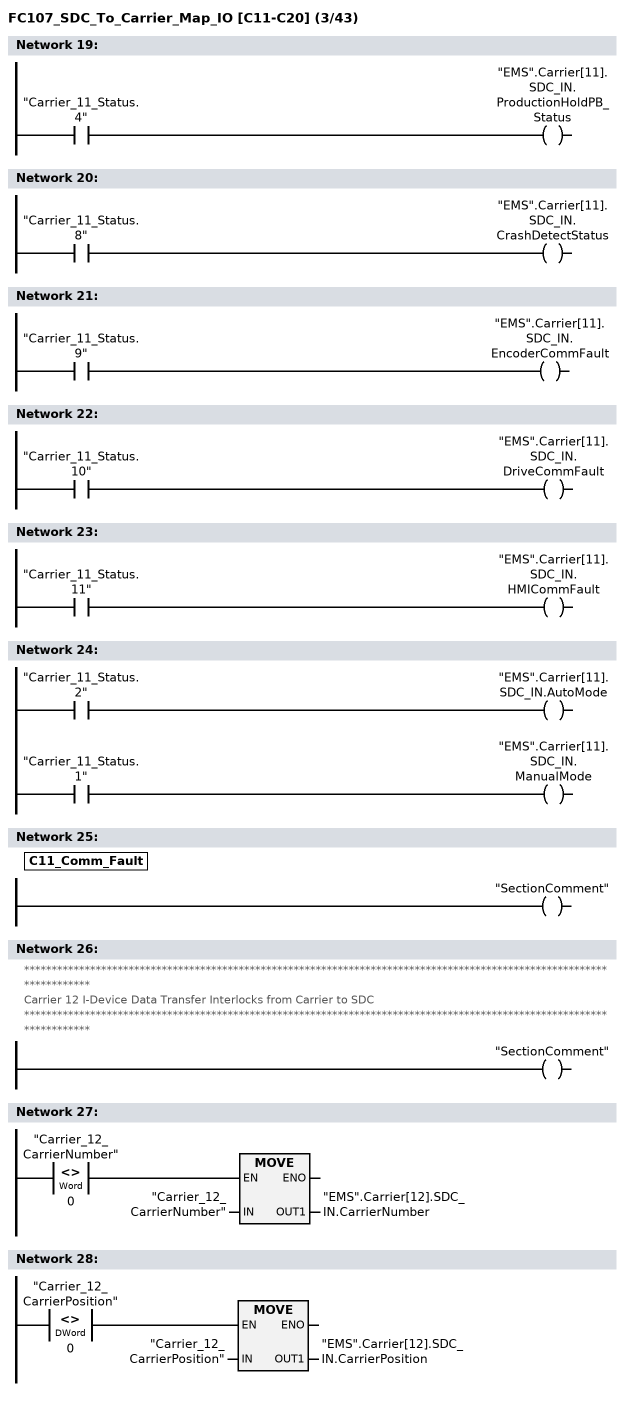
   RUNG wire#powerrail
      Contact( "Carrier_11_Status.4" )
      Coil( "EMS".Carrier[11].SDC_IN.ProductionHoldPB_Status )
   END_RUNG
   // the same network as SCL:
   "EMS".Carrier[11].SDC_IN.ProductionHoldPB_Status := "Carrier_11_Status.4";
END_REGION

REGION Network 20
   RUNG wire#powerrail
      Contact( "Carrier_11_Status.8" )
      Coil( "EMS".Carrier[11].SDC_IN.CrashDetectStatus )
   END_RUNG
   // the same network as SCL:
   "EMS".Carrier[11].SDC_IN.CrashDetectStatus := "Carrier_11_Status.8";
END_REGION

REGION Network 21
   RUNG wire#powerrail
      Contact( "Carrier_11_Status.9" )
      Coil( "EMS".Carrier[11].SDC_IN.EncoderCommFault )
   END_RUNG
   // the same network as SCL:
   "EMS".Carrier[11].SDC_IN.EncoderCommFault := "Carrier_11_Status.9";
END_REGION

REGION Network 22
   RUNG wire#powerrail
      Contact( "Carrier_11_Status.10" )
      Coil( "EMS".Carrier[11].SDC_IN.DriveCommFault )
   END_RUNG
   // the same network as SCL:
   "EMS".Carrier[11].SDC_IN.DriveCommFault := "Carrier_11_Status.10";
END_REGION

REGION Network 23
   RUNG wire#powerrail
      Contact( "Carrier_11_Status.11" )
      Coil( "EMS".Carrier[11].SDC_IN.HMICommFault )
   END_RUNG
   // the same network as SCL:
   "EMS".Carrier[11].SDC_IN.HMICommFault := "Carrier_11_Status.11";
END_REGION

REGION Network 24
   RUNG wire#powerrail
      Contact( "Carrier_11_Status.2" )
      Coil( "EMS".Carrier[11].SDC_IN.AutoMode )
   END_RUNG
   RUNG wire#powerrail
      Contact( "Carrier_11_Status.1" )
      Coil( "EMS".Carrier[11].SDC_IN.ManualMode )
   END_RUNG
   // the same network as SCL:
   "EMS".Carrier[11].SDC_IN.AutoMode := "Carrier_11_Status.2";
   "EMS".Carrier[11].SDC_IN.ManualMode := "Carrier_11_Status.1";
END_REGION

REGION Network 25
   Label( C11_Comm_Fault )
   RUNG wire#powerrail
      Coil( "SectionComment" )
   END_RUNG
   // the same network as SCL:
   C11_Comm_Fault:
   "SectionComment" := TRUE;
END_REGION

REGION Network 26
   // **********************************************************************************************************************
   // 
   // Carrier 12 I-Device Data Transfer Interlocks from Carrier to SDC
   // 
   // **********************************************************************************************************************
   RUNG wire#powerrail
      Coil( "SectionComment" )
   END_RUNG
   // the same network as SCL:
   "SectionComment" := TRUE;
END_REGION

REGION Network 27
   RUNG wire#powerrail
      { S7_Templates := "SrcType := Word" } NE_Contact(in1 := "Carrier_12_CarrierNumber", in2 := 0)
      Move(in := "Carrier_12_CarrierNumber", out1 => "EMS".Carrier[12].SDC_IN.CarrierNumber)
   END_RUNG
   // the same network as SCL:
   IF "Carrier_12_CarrierNumber" <> 0 THEN
       "EMS".Carrier[12].SDC_IN.CarrierNumber := "Carrier_12_CarrierNumber";
   END_IF;
END_REGION

REGION Network 28
   RUNG wire#powerrail
      { S7_Templates := "SrcType := DWord" } NE_Contact(in1 := "Carrier_12_CarrierPosition", in2 := 0)
      Move(in := "Carrier_12_CarrierPosition", out1 => "EMS".Carrier[12].SDC_IN.CarrierPosition)
   END_RUNG
   // the same network as SCL:
   IF "Carrier_12_CarrierPosition" <> 0 THEN
       "EMS".Carrier[12].SDC_IN.CarrierPosition := "Carrier_12_CarrierPosition";
   END_IF;
END_REGION

REGION Network 29
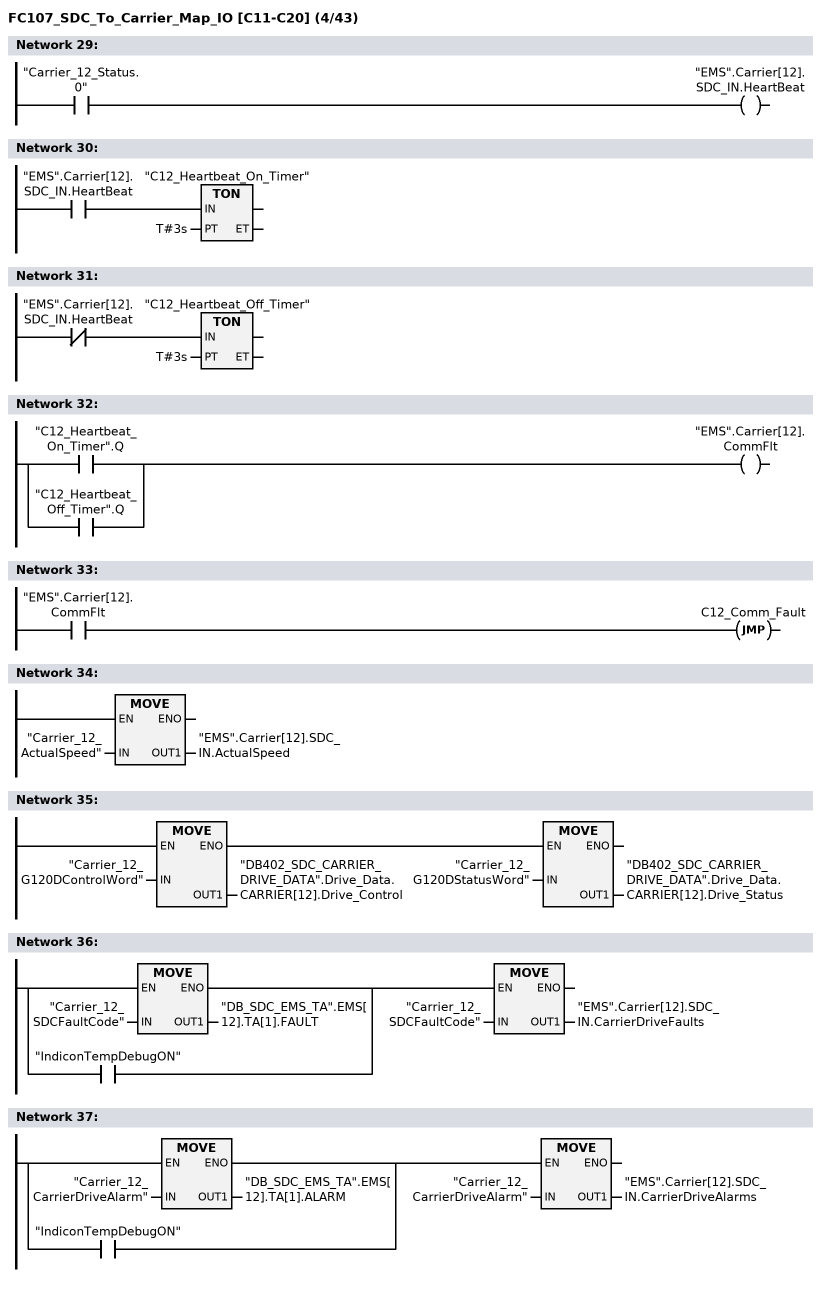
   RUNG wire#powerrail
      Contact( "Carrier_12_Status.0" )
      Coil( "EMS".Carrier[12].SDC_IN.HeartBeat )
   END_RUNG
   // the same network as SCL:
   "EMS".Carrier[12].SDC_IN.HeartBeat := "Carrier_12_Status.0";
END_REGION

REGION Network 30
   "C12_Heartbeat_On_Timer".TON(IN := "EMS".Carrier[12].SDC_IN.HeartBeat, PT := T#3s);
END_REGION

REGION Network 31
   "C12_Heartbeat_Off_Timer".TON(IN := NOT "EMS".Carrier[12].SDC_IN.HeartBeat, PT := T#3s);
END_REGION

REGION Network 32
   RUNG wire#powerrail
      Contact( "C12_Heartbeat_On_Timer".Q )
      wire#w1
      Coil( "EMS".Carrier[12].CommFlt )
   END_RUNG
   RUNG wire#powerrail
      Contact( "C12_Heartbeat_Off_Timer".Q )
   END_RUNG wire#w1
   // the same network as SCL:
   "EMS".Carrier[12].CommFlt := "C12_Heartbeat_On_Timer".Q OR "C12_Heartbeat_Off_Timer".Q;
END_REGION

REGION Network 33
   RUNG wire#powerrail
      Contact( "EMS".Carrier[12].CommFlt )
      JumpCoil( C12_Comm_Fault )
   END_RUNG
   // the same network as SCL:
   IF "EMS".Carrier[12].CommFlt THEN GOTO C12_Comm_Fault; END_IF;
END_REGION

REGION Network 34
   RUNG wire#powerrail
      Move(in := "Carrier_12_ActualSpeed", out1 => "EMS".Carrier[12].SDC_IN.ActualSpeed)
   END_RUNG
   // the same network as SCL:
   "EMS".Carrier[12].SDC_IN.ActualSpeed := "Carrier_12_ActualSpeed";
END_REGION

REGION Network 35
   RUNG wire#powerrail
      Move(in := "Carrier_12_G120DControlWord", out1 => "DB402_SDC_CARRIER_DRIVE_DATA".Drive_Data.CARRIER[12].Drive_Control)
      Move(in := "Carrier_12_G120DStatusWord", out1 => "DB402_SDC_CARRIER_DRIVE_DATA".Drive_Data.CARRIER[12].Drive_Status)
   END_RUNG
   // the same network as SCL:
   "DB402_SDC_CARRIER_DRIVE_DATA".Drive_Data.CARRIER[12].Drive_Control := "Carrier_12_G120DControlWord";
   "DB402_SDC_CARRIER_DRIVE_DATA".Drive_Data.CARRIER[12].Drive_Status := "Carrier_12_G120DStatusWord";
END_REGION

REGION Network 36
   RUNG wire#powerrail
      Move(in := "Carrier_12_SDCFaultCode", out1 => "DB_SDC_EMS_TA".EMS[12].TA[1].FAULT)
      wire#w1
      Move(in := "Carrier_12_SDCFaultCode", out1 => "EMS".Carrier[12].SDC_IN.CarrierDriveFaults)
   END_RUNG
   RUNG wire#powerrail
      Contact( "IndiconTempDebugON" )
   END_RUNG wire#w1
   // the same network as SCL:
   "DB_SDC_EMS_TA".EMS[12].TA[1].FAULT := "Carrier_12_SDCFaultCode";
   IF TRUE OR "IndiconTempDebugON" THEN
       "EMS".Carrier[12].SDC_IN.CarrierDriveFaults := "Carrier_12_SDCFaultCode";
   END_IF;
END_REGION

REGION Network 37
   RUNG wire#powerrail
      Move(in := "Carrier_12_CarrierDriveAlarm", out1 => "DB_SDC_EMS_TA".EMS[12].TA[1].ALARM)
      wire#w1
      Move(in := "Carrier_12_CarrierDriveAlarm", out1 => "EMS".Carrier[12].SDC_IN.CarrierDriveAlarms)
   END_RUNG
   RUNG wire#powerrail
      Contact( "IndiconTempDebugON" )
   END_RUNG wire#w1
   // the same network as SCL:
   "DB_SDC_EMS_TA".EMS[12].TA[1].ALARM := "Carrier_12_CarrierDriveAlarm";
   IF TRUE OR "IndiconTempDebugON" THEN
       "EMS".Carrier[12].SDC_IN.CarrierDriveAlarms := "Carrier_12_CarrierDriveAlarm";
   END_IF;
END_REGION

REGION Network 38
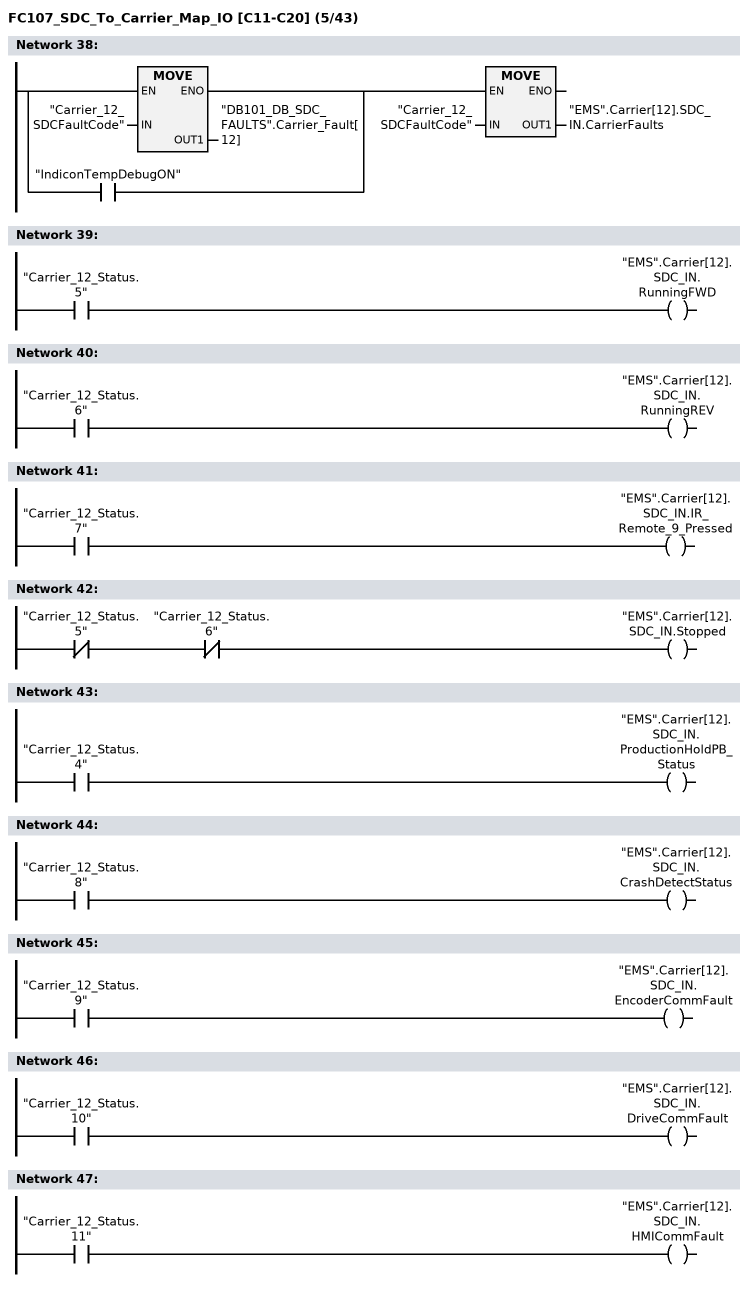
   RUNG wire#powerrail
      Move(in := "Carrier_12_SDCFaultCode", out1 => "DB101_DB_SDC_FAULTS".Carrier_Fault[12])
      wire#w1
      Move(in := "Carrier_12_SDCFaultCode", out1 => "EMS".Carrier[12].SDC_IN.CarrierFaults)
   END_RUNG
   RUNG wire#powerrail
      Contact( "IndiconTempDebugON" )
   END_RUNG wire#w1
   // the same network as SCL:
   "DB101_DB_SDC_FAULTS".Carrier_Fault[12] := "Carrier_12_SDCFaultCode";
   IF TRUE OR "IndiconTempDebugON" THEN
       "EMS".Carrier[12].SDC_IN.CarrierFaults := "Carrier_12_SDCFaultCode";
   END_IF;
END_REGION

REGION Network 39
   RUNG wire#powerrail
      Contact( "Carrier_12_Status.5" )
      Coil( "EMS".Carrier[12].SDC_IN.RunningFWD )
   END_RUNG
   // the same network as SCL:
   "EMS".Carrier[12].SDC_IN.RunningFWD := "Carrier_12_Status.5";
END_REGION

REGION Network 40
   RUNG wire#powerrail
      Contact( "Carrier_12_Status.6" )
      Coil( "EMS".Carrier[12].SDC_IN.RunningREV )
   END_RUNG
   // the same network as SCL:
   "EMS".Carrier[12].SDC_IN.RunningREV := "Carrier_12_Status.6";
END_REGION

REGION Network 41
   RUNG wire#powerrail
      Contact( "Carrier_12_Status.7" )
      Coil( "EMS".Carrier[12].SDC_IN.IR_Remote_9_Pressed )
   END_RUNG
   // the same network as SCL:
   "EMS".Carrier[12].SDC_IN.IR_Remote_9_Pressed := "Carrier_12_Status.7";
END_REGION

REGION Network 42
   RUNG wire#powerrail
      I_Contact( "Carrier_12_Status.5" )
      I_Contact( "Carrier_12_Status.6" )
      Coil( "EMS".Carrier[12].SDC_IN.Stopped )
   END_RUNG
   // the same network as SCL:
   "EMS".Carrier[12].SDC_IN.Stopped := NOT "Carrier_12_Status.5" AND NOT "Carrier_12_Status.6";
END_REGION

REGION Network 43
   RUNG wire#powerrail
      Contact( "Carrier_12_Status.4" )
      Coil( "EMS".Carrier[12].SDC_IN.ProductionHoldPB_Status )
   END_RUNG
   // the same network as SCL:
   "EMS".Carrier[12].SDC_IN.ProductionHoldPB_Status := "Carrier_12_Status.4";
END_REGION

REGION Network 44
   RUNG wire#powerrail
      Contact( "Carrier_12_Status.8" )
      Coil( "EMS".Carrier[12].SDC_IN.CrashDetectStatus )
   END_RUNG
   // the same network as SCL:
   "EMS".Carrier[12].SDC_IN.CrashDetectStatus := "Carrier_12_Status.8";
END_REGION

REGION Network 45
   RUNG wire#powerrail
      Contact( "Carrier_12_Status.9" )
      Coil( "EMS".Carrier[12].SDC_IN.EncoderCommFault )
   END_RUNG
   // the same network as SCL:
   "EMS".Carrier[12].SDC_IN.EncoderCommFault := "Carrier_12_Status.9";
END_REGION

REGION Network 46
   RUNG wire#powerrail
      Contact( "Carrier_12_Status.10" )
      Coil( "EMS".Carrier[12].SDC_IN.DriveCommFault )
   END_RUNG
   // the same network as SCL:
   "EMS".Carrier[12].SDC_IN.DriveCommFault := "Carrier_12_Status.10";
END_REGION

REGION Network 47
   RUNG wire#powerrail
      Contact( "Carrier_12_Status.11" )
      Coil( "EMS".Carrier[12].SDC_IN.HMICommFault )
   END_RUNG
   // the same network as SCL:
   "EMS".Carrier[12].SDC_IN.HMICommFault := "Carrier_12_Status.11";
END_REGION

REGION Network 48
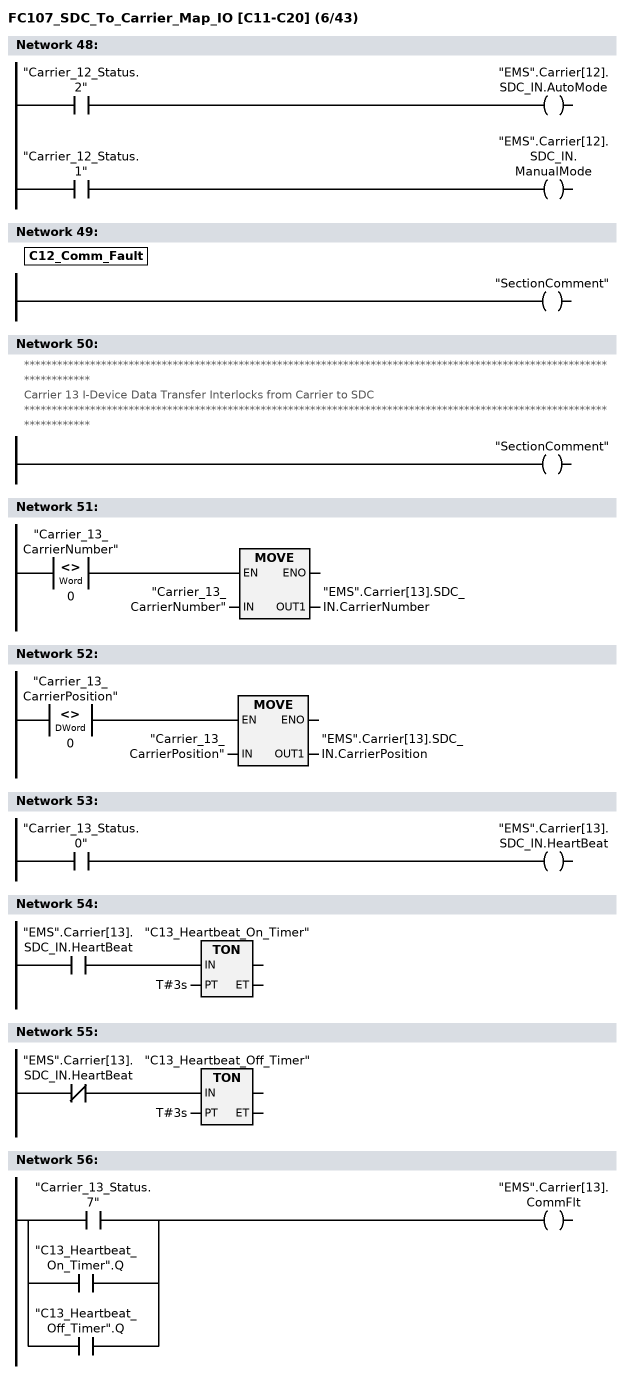
   RUNG wire#powerrail
      Contact( "Carrier_12_Status.2" )
      Coil( "EMS".Carrier[12].SDC_IN.AutoMode )
   END_RUNG
   RUNG wire#powerrail
      Contact( "Carrier_12_Status.1" )
      Coil( "EMS".Carrier[12].SDC_IN.ManualMode )
   END_RUNG
   // the same network as SCL:
   "EMS".Carrier[12].SDC_IN.AutoMode := "Carrier_12_Status.2";
   "EMS".Carrier[12].SDC_IN.ManualMode := "Carrier_12_Status.1";
END_REGION

REGION Network 49
   Label( C12_Comm_Fault )
   RUNG wire#powerrail
      Coil( "SectionComment" )
   END_RUNG
   // the same network as SCL:
   C12_Comm_Fault:
   "SectionComment" := TRUE;
END_REGION

REGION Network 50
   // **********************************************************************************************************************
   // 
   // Carrier 13 I-Device Data Transfer Interlocks from Carrier to SDC
   // 
   // **********************************************************************************************************************
   RUNG wire#powerrail
      Coil( "SectionComment" )
   END_RUNG
   // the same network as SCL:
   "SectionComment" := TRUE;
END_REGION

REGION Network 51
   RUNG wire#powerrail
      { S7_Templates := "SrcType := Word" } NE_Contact(in1 := "Carrier_13_CarrierNumber", in2 := 0)
      Move(in := "Carrier_13_CarrierNumber", out1 => "EMS".Carrier[13].SDC_IN.CarrierNumber)
   END_RUNG
   // the same network as SCL:
   IF "Carrier_13_CarrierNumber" <> 0 THEN
       "EMS".Carrier[13].SDC_IN.CarrierNumber := "Carrier_13_CarrierNumber";
   END_IF;
END_REGION

REGION Network 52
   RUNG wire#powerrail
      { S7_Templates := "SrcType := DWord" } NE_Contact(in1 := "Carrier_13_CarrierPosition", in2 := 0)
      Move(in := "Carrier_13_CarrierPosition", out1 => "EMS".Carrier[13].SDC_IN.CarrierPosition)
   END_RUNG
   // the same network as SCL:
   IF "Carrier_13_CarrierPosition" <> 0 THEN
       "EMS".Carrier[13].SDC_IN.CarrierPosition := "Carrier_13_CarrierPosition";
   END_IF;
END_REGION

REGION Network 53
   RUNG wire#powerrail
      Contact( "Carrier_13_Status.0" )
      Coil( "EMS".Carrier[13].SDC_IN.HeartBeat )
   END_RUNG
   // the same network as SCL:
   "EMS".Carrier[13].SDC_IN.HeartBeat := "Carrier_13_Status.0";
END_REGION

REGION Network 54
   "C13_Heartbeat_On_Timer".TON(IN := "EMS".Carrier[13].SDC_IN.HeartBeat, PT := T#3s);
END_REGION

REGION Network 55
   "C13_Heartbeat_Off_Timer".TON(IN := NOT "EMS".Carrier[13].SDC_IN.HeartBeat, PT := T#3s);
END_REGION

REGION Network 56
   RUNG wire#powerrail
      Contact( "Carrier_13_Status.7" )
      wire#w1
      Coil( "EMS".Carrier[13].CommFlt )
   END_RUNG
   RUNG wire#powerrail
      Contact( "C13_Heartbeat_On_Timer".Q )
   END_RUNG wire#w1
   RUNG wire#powerrail
      Contact( "C13_Heartbeat_Off_Timer".Q )
   END_RUNG wire#w1
   // the same network as SCL:
   "EMS".Carrier[13].CommFlt := "Carrier_13_Status.7" OR "C13_Heartbeat_On_Timer".Q OR "C13_Heartbeat_Off_Timer".Q;
END_REGION

REGION Network 57
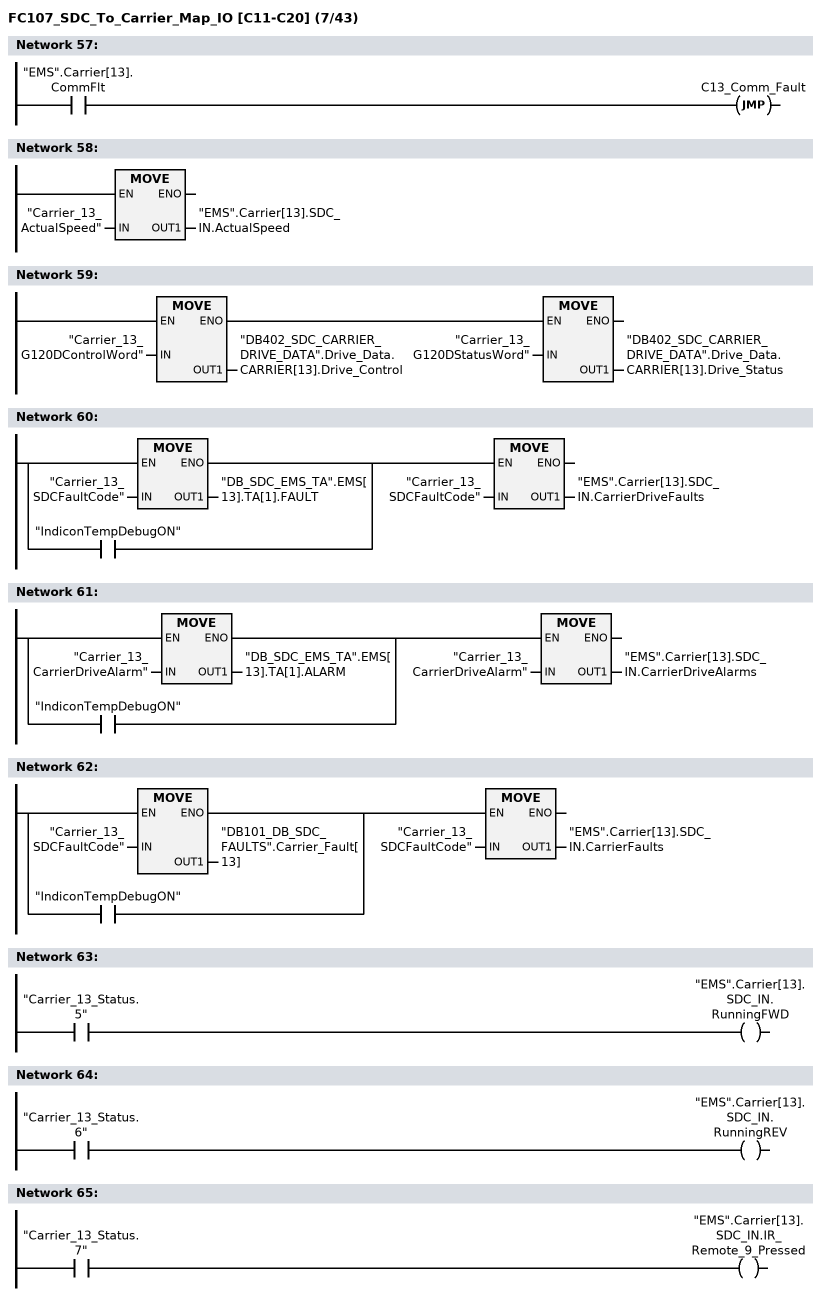
   RUNG wire#powerrail
      Contact( "EMS".Carrier[13].CommFlt )
      JumpCoil( C13_Comm_Fault )
   END_RUNG
   // the same network as SCL:
   IF "EMS".Carrier[13].CommFlt THEN GOTO C13_Comm_Fault; END_IF;
END_REGION

REGION Network 58
   RUNG wire#powerrail
      Move(in := "Carrier_13_ActualSpeed", out1 => "EMS".Carrier[13].SDC_IN.ActualSpeed)
   END_RUNG
   // the same network as SCL:
   "EMS".Carrier[13].SDC_IN.ActualSpeed := "Carrier_13_ActualSpeed";
END_REGION

REGION Network 59
   RUNG wire#powerrail
      Move(in := "Carrier_13_G120DControlWord", out1 => "DB402_SDC_CARRIER_DRIVE_DATA".Drive_Data.CARRIER[13].Drive_Control)
      Move(in := "Carrier_13_G120DStatusWord", out1 => "DB402_SDC_CARRIER_DRIVE_DATA".Drive_Data.CARRIER[13].Drive_Status)
   END_RUNG
   // the same network as SCL:
   "DB402_SDC_CARRIER_DRIVE_DATA".Drive_Data.CARRIER[13].Drive_Control := "Carrier_13_G120DControlWord";
   "DB402_SDC_CARRIER_DRIVE_DATA".Drive_Data.CARRIER[13].Drive_Status := "Carrier_13_G120DStatusWord";
END_REGION

REGION Network 60
   RUNG wire#powerrail
      Move(in := "Carrier_13_SDCFaultCode", out1 => "DB_SDC_EMS_TA".EMS[13].TA[1].FAULT)
      wire#w1
      Move(in := "Carrier_13_SDCFaultCode", out1 => "EMS".Carrier[13].SDC_IN.CarrierDriveFaults)
   END_RUNG
   RUNG wire#powerrail
      Contact( "IndiconTempDebugON" )
   END_RUNG wire#w1
   // the same network as SCL:
   "DB_SDC_EMS_TA".EMS[13].TA[1].FAULT := "Carrier_13_SDCFaultCode";
   IF TRUE OR "IndiconTempDebugON" THEN
       "EMS".Carrier[13].SDC_IN.CarrierDriveFaults := "Carrier_13_SDCFaultCode";
   END_IF;
END_REGION

REGION Network 61
   RUNG wire#powerrail
      Move(in := "Carrier_13_CarrierDriveAlarm", out1 => "DB_SDC_EMS_TA".EMS[13].TA[1].ALARM)
      wire#w1
      Move(in := "Carrier_13_CarrierDriveAlarm", out1 => "EMS".Carrier[13].SDC_IN.CarrierDriveAlarms)
   END_RUNG
   RUNG wire#powerrail
      Contact( "IndiconTempDebugON" )
   END_RUNG wire#w1
   // the same network as SCL:
   "DB_SDC_EMS_TA".EMS[13].TA[1].ALARM := "Carrier_13_CarrierDriveAlarm";
   IF TRUE OR "IndiconTempDebugON" THEN
       "EMS".Carrier[13].SDC_IN.CarrierDriveAlarms := "Carrier_13_CarrierDriveAlarm";
   END_IF;
END_REGION

REGION Network 62
   RUNG wire#powerrail
      Move(in := "Carrier_13_SDCFaultCode", out1 => "DB101_DB_SDC_FAULTS".Carrier_Fault[13])
      wire#w1
      Move(in := "Carrier_13_SDCFaultCode", out1 => "EMS".Carrier[13].SDC_IN.CarrierFaults)
   END_RUNG
   RUNG wire#powerrail
      Contact( "IndiconTempDebugON" )
   END_RUNG wire#w1
   // the same network as SCL:
   "DB101_DB_SDC_FAULTS".Carrier_Fault[13] := "Carrier_13_SDCFaultCode";
   IF TRUE OR "IndiconTempDebugON" THEN
       "EMS".Carrier[13].SDC_IN.CarrierFaults := "Carrier_13_SDCFaultCode";
   END_IF;
END_REGION

REGION Network 63
   RUNG wire#powerrail
      Contact( "Carrier_13_Status.5" )
      Coil( "EMS".Carrier[13].SDC_IN.RunningFWD )
   END_RUNG
   // the same network as SCL:
   "EMS".Carrier[13].SDC_IN.RunningFWD := "Carrier_13_Status.5";
END_REGION

REGION Network 64
   RUNG wire#powerrail
      Contact( "Carrier_13_Status.6" )
      Coil( "EMS".Carrier[13].SDC_IN.RunningREV )
   END_RUNG
   // the same network as SCL:
   "EMS".Carrier[13].SDC_IN.RunningREV := "Carrier_13_Status.6";
END_REGION

REGION Network 65
   RUNG wire#powerrail
      Contact( "Carrier_13_Status.7" )
      Coil( "EMS".Carrier[13].SDC_IN.IR_Remote_9_Pressed )
   END_RUNG
   // the same network as SCL:
   "EMS".Carrier[13].SDC_IN.IR_Remote_9_Pressed := "Carrier_13_Status.7";
END_REGION

REGION Network 66
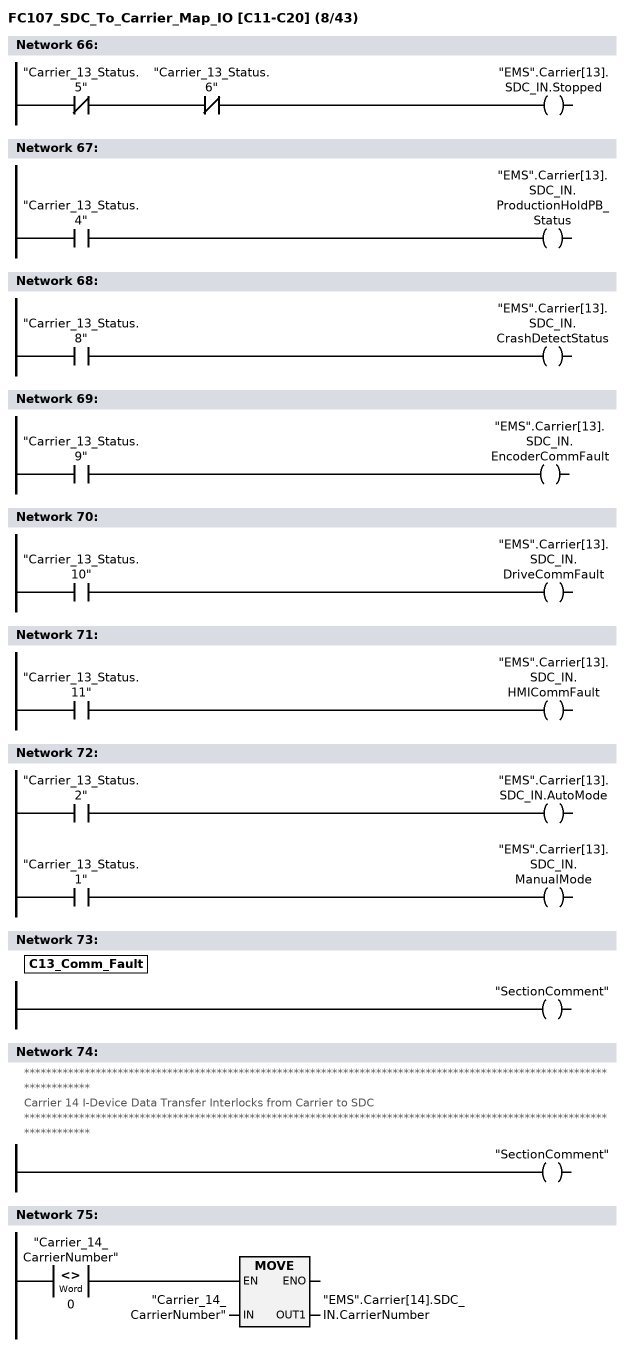
   RUNG wire#powerrail
      I_Contact( "Carrier_13_Status.5" )
      I_Contact( "Carrier_13_Status.6" )
      Coil( "EMS".Carrier[13].SDC_IN.Stopped )
   END_RUNG
   // the same network as SCL:
   "EMS".Carrier[13].SDC_IN.Stopped := NOT "Carrier_13_Status.5" AND NOT "Carrier_13_Status.6";
END_REGION

REGION Network 67
   RUNG wire#powerrail
      Contact( "Carrier_13_Status.4" )
      Coil( "EMS".Carrier[13].SDC_IN.ProductionHoldPB_Status )
   END_RUNG
   // the same network as SCL:
   "EMS".Carrier[13].SDC_IN.ProductionHoldPB_Status := "Carrier_13_Status.4";
END_REGION

REGION Network 68
   RUNG wire#powerrail
      Contact( "Carrier_13_Status.8" )
      Coil( "EMS".Carrier[13].SDC_IN.CrashDetectStatus )
   END_RUNG
   // the same network as SCL:
   "EMS".Carrier[13].SDC_IN.CrashDetectStatus := "Carrier_13_Status.8";
END_REGION

REGION Network 69
   RUNG wire#powerrail
      Contact( "Carrier_13_Status.9" )
      Coil( "EMS".Carrier[13].SDC_IN.EncoderCommFault )
   END_RUNG
   // the same network as SCL:
   "EMS".Carrier[13].SDC_IN.EncoderCommFault := "Carrier_13_Status.9";
END_REGION

REGION Network 70
   RUNG wire#powerrail
      Contact( "Carrier_13_Status.10" )
      Coil( "EMS".Carrier[13].SDC_IN.DriveCommFault )
   END_RUNG
   // the same network as SCL:
   "EMS".Carrier[13].SDC_IN.DriveCommFault := "Carrier_13_Status.10";
END_REGION

REGION Network 71
   RUNG wire#powerrail
      Contact( "Carrier_13_Status.11" )
      Coil( "EMS".Carrier[13].SDC_IN.HMICommFault )
   END_RUNG
   // the same network as SCL:
   "EMS".Carrier[13].SDC_IN.HMICommFault := "Carrier_13_Status.11";
END_REGION

REGION Network 72
   RUNG wire#powerrail
      Contact( "Carrier_13_Status.2" )
      Coil( "EMS".Carrier[13].SDC_IN.AutoMode )
   END_RUNG
   RUNG wire#powerrail
      Contact( "Carrier_13_Status.1" )
      Coil( "EMS".Carrier[13].SDC_IN.ManualMode )
   END_RUNG
   // the same network as SCL:
   "EMS".Carrier[13].SDC_IN.AutoMode := "Carrier_13_Status.2";
   "EMS".Carrier[13].SDC_IN.ManualMode := "Carrier_13_Status.1";
END_REGION

REGION Network 73
   Label( C13_Comm_Fault )
   RUNG wire#powerrail
      Coil( "SectionComment" )
   END_RUNG
   // the same network as SCL:
   C13_Comm_Fault:
   "SectionComment" := TRUE;
END_REGION

REGION Network 74
   // **********************************************************************************************************************
   // 
   // Carrier 14 I-Device Data Transfer Interlocks from Carrier to SDC
   // 
   // **********************************************************************************************************************
   RUNG wire#powerrail
      Coil( "SectionComment" )
   END_RUNG
   // the same network as SCL:
   "SectionComment" := TRUE;
END_REGION

REGION Network 75
   RUNG wire#powerrail
      { S7_Templates := "SrcType := Word" } NE_Contact(in1 := "Carrier_14_CarrierNumber", in2 := 0)
      Move(in := "Carrier_14_CarrierNumber", out1 => "EMS".Carrier[14].SDC_IN.CarrierNumber)
   END_RUNG
   // the same network as SCL:
   IF "Carrier_14_CarrierNumber" <> 0 THEN
       "EMS".Carrier[14].SDC_IN.CarrierNumber := "Carrier_14_CarrierNumber";
   END_IF;
END_REGION

REGION Network 76
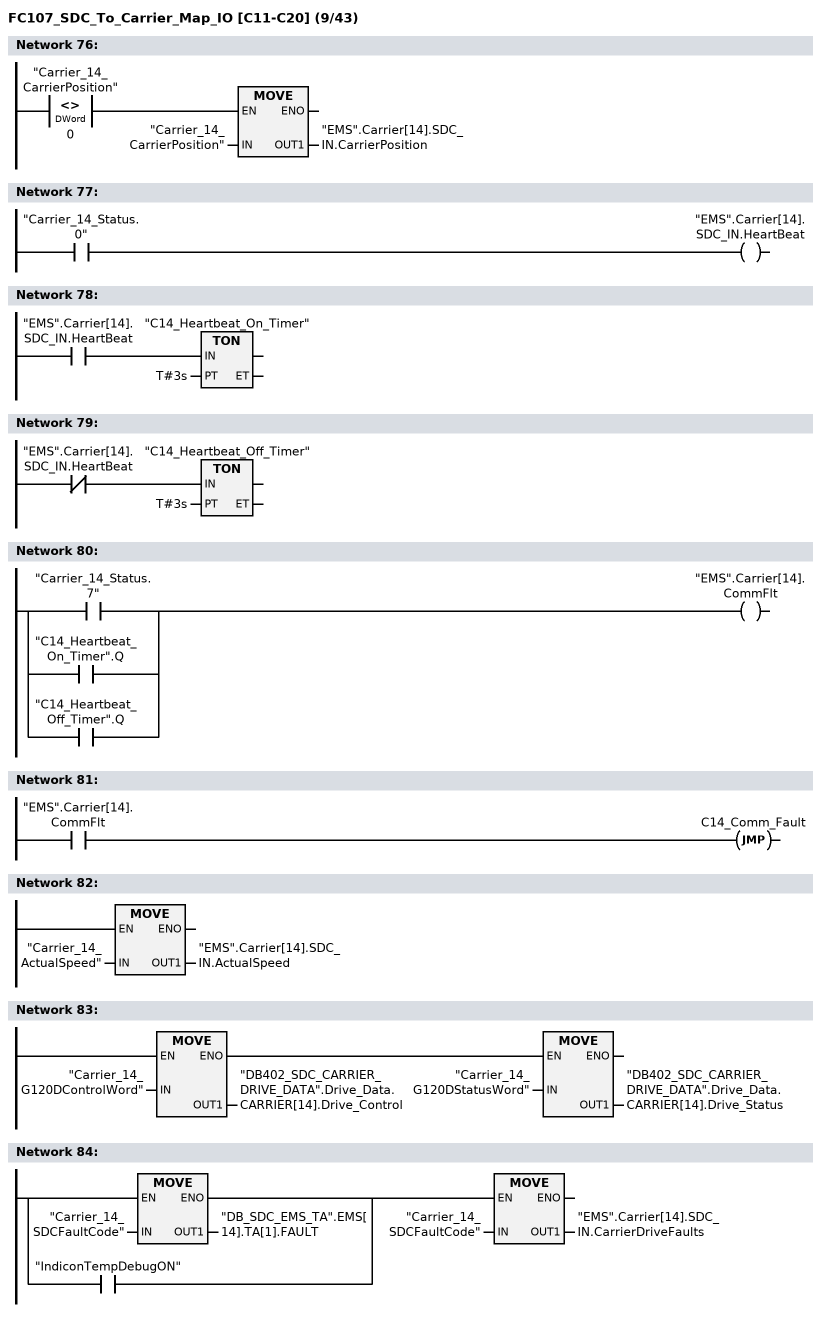
   RUNG wire#powerrail
      { S7_Templates := "SrcType := DWord" } NE_Contact(in1 := "Carrier_14_CarrierPosition", in2 := 0)
      Move(in := "Carrier_14_CarrierPosition", out1 => "EMS".Carrier[14].SDC_IN.CarrierPosition)
   END_RUNG
   // the same network as SCL:
   IF "Carrier_14_CarrierPosition" <> 0 THEN
       "EMS".Carrier[14].SDC_IN.CarrierPosition := "Carrier_14_CarrierPosition";
   END_IF;
END_REGION

REGION Network 77
   RUNG wire#powerrail
      Contact( "Carrier_14_Status.0" )
      Coil( "EMS".Carrier[14].SDC_IN.HeartBeat )
   END_RUNG
   // the same network as SCL:
   "EMS".Carrier[14].SDC_IN.HeartBeat := "Carrier_14_Status.0";
END_REGION

REGION Network 78
   "C14_Heartbeat_On_Timer".TON(IN := "EMS".Carrier[14].SDC_IN.HeartBeat, PT := T#3s);
END_REGION

REGION Network 79
   "C14_Heartbeat_Off_Timer".TON(IN := NOT "EMS".Carrier[14].SDC_IN.HeartBeat, PT := T#3s);
END_REGION

REGION Network 80
   RUNG wire#powerrail
      Contact( "Carrier_14_Status.7" )
      wire#w1
      Coil( "EMS".Carrier[14].CommFlt )
   END_RUNG
   RUNG wire#powerrail
      Contact( "C14_Heartbeat_On_Timer".Q )
   END_RUNG wire#w1
   RUNG wire#powerrail
      Contact( "C14_Heartbeat_Off_Timer".Q )
   END_RUNG wire#w1
   // the same network as SCL:
   "EMS".Carrier[14].CommFlt := "Carrier_14_Status.7" OR "C14_Heartbeat_On_Timer".Q OR "C14_Heartbeat_Off_Timer".Q;
END_REGION

REGION Network 81
   RUNG wire#powerrail
      Contact( "EMS".Carrier[14].CommFlt )
      JumpCoil( C14_Comm_Fault )
   END_RUNG
   // the same network as SCL:
   IF "EMS".Carrier[14].CommFlt THEN GOTO C14_Comm_Fault; END_IF;
END_REGION

REGION Network 82
   RUNG wire#powerrail
      Move(in := "Carrier_14_ActualSpeed", out1 => "EMS".Carrier[14].SDC_IN.ActualSpeed)
   END_RUNG
   // the same network as SCL:
   "EMS".Carrier[14].SDC_IN.ActualSpeed := "Carrier_14_ActualSpeed";
END_REGION

REGION Network 83
   RUNG wire#powerrail
      Move(in := "Carrier_14_G120DControlWord", out1 => "DB402_SDC_CARRIER_DRIVE_DATA".Drive_Data.CARRIER[14].Drive_Control)
      Move(in := "Carrier_14_G120DStatusWord", out1 => "DB402_SDC_CARRIER_DRIVE_DATA".Drive_Data.CARRIER[14].Drive_Status)
   END_RUNG
   // the same network as SCL:
   "DB402_SDC_CARRIER_DRIVE_DATA".Drive_Data.CARRIER[14].Drive_Control := "Carrier_14_G120DControlWord";
   "DB402_SDC_CARRIER_DRIVE_DATA".Drive_Data.CARRIER[14].Drive_Status := "Carrier_14_G120DStatusWord";
END_REGION

REGION Network 84
   RUNG wire#powerrail
      Move(in := "Carrier_14_SDCFaultCode", out1 => "DB_SDC_EMS_TA".EMS[14].TA[1].FAULT)
      wire#w1
      Move(in := "Carrier_14_SDCFaultCode", out1 => "EMS".Carrier[14].SDC_IN.CarrierDriveFaults)
   END_RUNG
   RUNG wire#powerrail
      Contact( "IndiconTempDebugON" )
   END_RUNG wire#w1
   // the same network as SCL:
   "DB_SDC_EMS_TA".EMS[14].TA[1].FAULT := "Carrier_14_SDCFaultCode";
   IF TRUE OR "IndiconTempDebugON" THEN
       "EMS".Carrier[14].SDC_IN.CarrierDriveFaults := "Carrier_14_SDCFaultCode";
   END_IF;
END_REGION

REGION Network 85
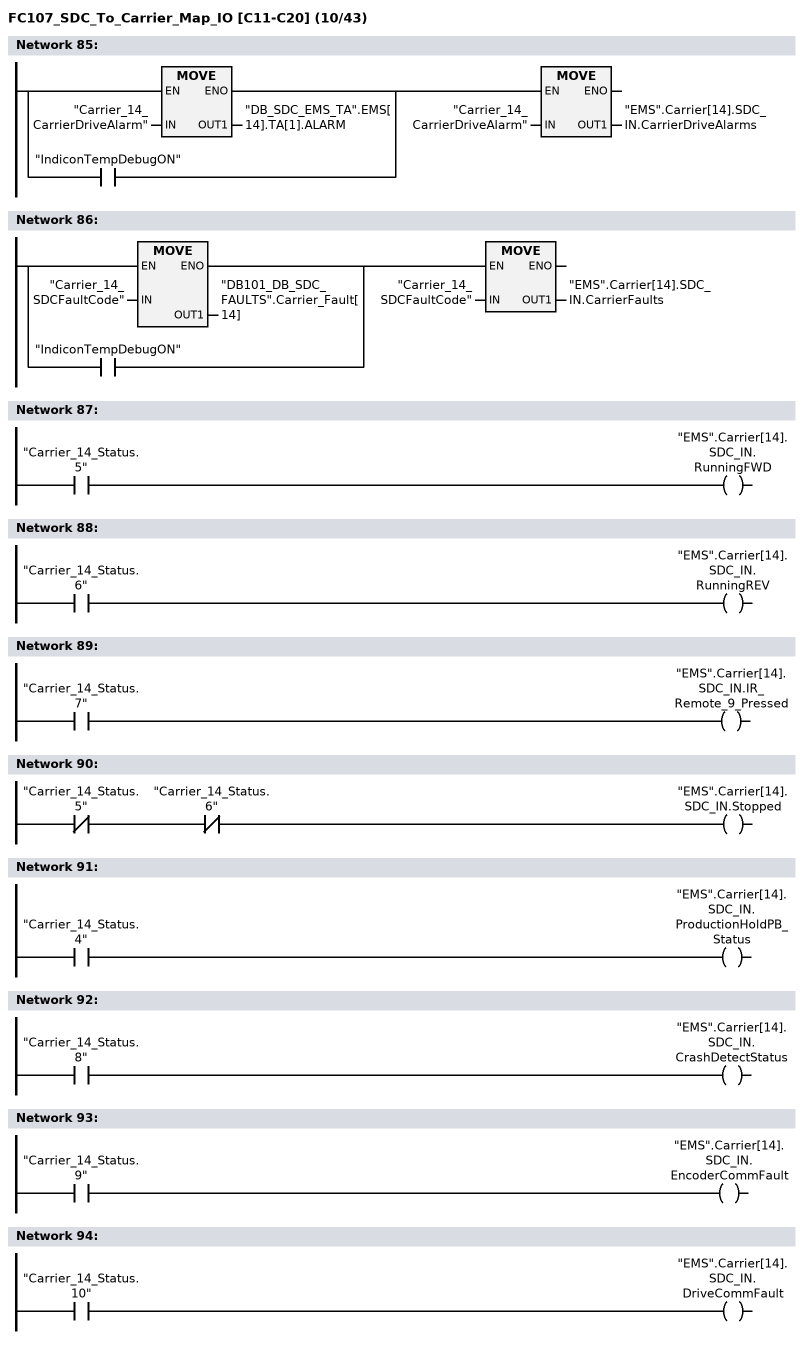
   RUNG wire#powerrail
      Move(in := "Carrier_14_CarrierDriveAlarm", out1 => "DB_SDC_EMS_TA".EMS[14].TA[1].ALARM)
      wire#w1
      Move(in := "Carrier_14_CarrierDriveAlarm", out1 => "EMS".Carrier[14].SDC_IN.CarrierDriveAlarms)
   END_RUNG
   RUNG wire#powerrail
      Contact( "IndiconTempDebugON" )
   END_RUNG wire#w1
   // the same network as SCL:
   "DB_SDC_EMS_TA".EMS[14].TA[1].ALARM := "Carrier_14_CarrierDriveAlarm";
   IF TRUE OR "IndiconTempDebugON" THEN
       "EMS".Carrier[14].SDC_IN.CarrierDriveAlarms := "Carrier_14_CarrierDriveAlarm";
   END_IF;
END_REGION

REGION Network 86
   RUNG wire#powerrail
      Move(in := "Carrier_14_SDCFaultCode", out1 => "DB101_DB_SDC_FAULTS".Carrier_Fault[14])
      wire#w1
      Move(in := "Carrier_14_SDCFaultCode", out1 => "EMS".Carrier[14].SDC_IN.CarrierFaults)
   END_RUNG
   RUNG wire#powerrail
      Contact( "IndiconTempDebugON" )
   END_RUNG wire#w1
   // the same network as SCL:
   "DB101_DB_SDC_FAULTS".Carrier_Fault[14] := "Carrier_14_SDCFaultCode";
   IF TRUE OR "IndiconTempDebugON" THEN
       "EMS".Carrier[14].SDC_IN.CarrierFaults := "Carrier_14_SDCFaultCode";
   END_IF;
END_REGION

REGION Network 87
   RUNG wire#powerrail
      Contact( "Carrier_14_Status.5" )
      Coil( "EMS".Carrier[14].SDC_IN.RunningFWD )
   END_RUNG
   // the same network as SCL:
   "EMS".Carrier[14].SDC_IN.RunningFWD := "Carrier_14_Status.5";
END_REGION

REGION Network 88
   RUNG wire#powerrail
      Contact( "Carrier_14_Status.6" )
      Coil( "EMS".Carrier[14].SDC_IN.RunningREV )
   END_RUNG
   // the same network as SCL:
   "EMS".Carrier[14].SDC_IN.RunningREV := "Carrier_14_Status.6";
END_REGION

REGION Network 89
   RUNG wire#powerrail
      Contact( "Carrier_14_Status.7" )
      Coil( "EMS".Carrier[14].SDC_IN.IR_Remote_9_Pressed )
   END_RUNG
   // the same network as SCL:
   "EMS".Carrier[14].SDC_IN.IR_Remote_9_Pressed := "Carrier_14_Status.7";
END_REGION

REGION Network 90
   RUNG wire#powerrail
      I_Contact( "Carrier_14_Status.5" )
      I_Contact( "Carrier_14_Status.6" )
      Coil( "EMS".Carrier[14].SDC_IN.Stopped )
   END_RUNG
   // the same network as SCL:
   "EMS".Carrier[14].SDC_IN.Stopped := NOT "Carrier_14_Status.5" AND NOT "Carrier_14_Status.6";
END_REGION

REGION Network 91
   RUNG wire#powerrail
      Contact( "Carrier_14_Status.4" )
      Coil( "EMS".Carrier[14].SDC_IN.ProductionHoldPB_Status )
   END_RUNG
   // the same network as SCL:
   "EMS".Carrier[14].SDC_IN.ProductionHoldPB_Status := "Carrier_14_Status.4";
END_REGION
